screen "Proses" 800x480, template "Template_1"
   TextField "Text field_18" at 473,92 size 53x19; Text 'TT-0001'
   IOField "I/O field_11" at 473,110 size 55x20; FormatPattern 999; Unit  °C
      ProcessValue <- "TT-0001"
   TextField "Text field_19" at 548,92 size 53x19; Text 'TT-0002'
   IOField "I/O field_12" at 548,110 size 55x20; FormatPattern 999; Unit  °C
      ProcessValue <- "TT-0002"
   TextField "Text field_20" at 474,141 size 50x19; Text 'PT-0001'
   IOField "I/O field_13" at 474,159 size 52x20; FormatPattern 99; Unit  Bar
      ProcessValue <- "PT-0001"
   TextField "Text field_21" at 550,141 size 50x19; Text 'PT-0002'
   IOField "I/O field_14" at 550,159 size 52x20; FormatPattern 99; Unit  Bar
      ProcessValue <- "PT-0002"
   GraphicView "Graphic view_17" at 37,119 size 60x45; Picture "Graphic_29"
   Circle "Circle_3" at 95,98 size 16x16
      Appearance <- "PUMP_PUMP-1_Yedek1"
   TextField "Text field_67" at 24,118 size 16x22; Text 'R'
      Visibility <- "PUMP_PUMP-1_Local/Remote"
   TextField "Text field_68" at 26,119 size 14x22; Text 'L'
      Visibility <- "PUMP_PUMP-1_Local/Remote"
   TextField "Text field_10" at 28,97 size 49x20; Text 'PUMP-1'
   IOField "I/O field_15" at 71,167 size 45x20; FormatPattern 99; Unit  A
      ProcessValue <- "Pump-1_A"
   IOField "I/O field_6" at 24,167 size 45x20; FormatPattern 999; Unit  °C
      ProcessValue <- "Pump-1_Temp"
   GraphicView "Graphic view_1" at 145,119 size 60x45; Picture "Graphic_29"
   Circle "Circle_1" at 203,98 size 16x16
      Appearance <- "PUMP_PUMP-2_Yedek1"
   TextField "Text field_1" at 132,118 size 16x22; Text 'R'
      Visibility <- "PUMP_PUMP-2_Local/Remote"
   TextField "Text field_2" at 134,117 size 14x22; Text 'L'
      Visibility <- "PUMP_PUMP-2_Local/Remote"
   TextField "Text field_3" at 136,97 size 49x20; Text 'PUMP-2'
   IOField "I/O field_1" at 179,167 size 45x20; FormatPattern 99; Unit  A
      ProcessValue <- "Pump-2_A"
   IOField "I/O field_2" at 132,167 size 45x20; FormatPattern 999; Unit  °C
      ProcessValue <- "Pump-2_Temp"
   GraphicView "Graphic view_2" at 254,119 size 60x45; Picture "Graphic_29"
   Circle "Circle_2" at 312,98 size 16x16
      Appearance <- "PUMP_PUMP-3_Yedek1"
   TextField "Text field_4" at 241,118 size 16x22; Text 'R'
      Visibility <- "PUMP_PUMP-3_Local/Remote"
   TextField "Text field_5" at 243,117 size 14x22; Text 'L'
      Visibility <- "PUMP_PUMP-3_Local/Remote"
   TextField "Text field_6" at 245,97 size 49x20; Text 'PUMP-3'
   IOField "I/O field_3" at 288,167 size 45x20; FormatPattern 99; Unit  A
      ProcessValue <- "Pump-3_A"
   IOField "I/O field_4" at 241,167 size 45x20; FormatPattern 999; Unit  °C
      ProcessValue <- "Pump-3_Temp"
   GraphicView "Graphic view_3" at 360,119 size 60x45; Picture "Graphic_29"
   Circle "Circle_4" at 418,98 size 16x16
      Appearance <- "PUMP_PUMP-4_Yedek1"
   TextField "Text field_7" at 347,118 size 16x22; Text 'R'
      Visibility <- "PUMP_PUMP-4_Local/Remote"
   TextField "Text field_8" at 349,117 size 14x22; Text 'L'
      Visibility <- "PUMP_PUMP-4_Local/Remote"
   TextField "Text field_9" at 351,97 size 49x20; Text 'PUMP-4'
   IOField "I/O field_5" at 394,167 size 45x20; FormatPattern 99; Unit  A
      ProcessValue <- "Pump-4_A"
   IOField "I/O field_7" at 347,167 size 45x20; FormatPattern 999; Unit  °C
      ProcessValue <- "Pump-4_Temp"
   IOField "I/O field_22" at 40,269 size 51x20; FormatPattern 9999; Unit  %
      ProcessValue <- "CValve-1_Fbk"
   TextField "Text field_70" at 32,212 size 74x19; Text 'CONTROL V-1'
   GraphicView "Template_Graphic view_5" at 44,232 size 38x32; Picture "Graphic_74"
   IOField "I/O field_8" at 148,269 size 51x20; FormatPattern 9999; Unit  %
      ProcessValue <- "CValve-2_Fbk"
   GraphicView "Template_Graphic view_1" at 152,232 size 38x32; Picture "Graphic_74"
   TextField "Text field_12" at 140,212 size 74x19; Text 'CONTROL V-2'
   IOField "I/O field_9" at 257,269 size 51x20; FormatPattern 9999; Unit  %
      ProcessValue <- "CValve-3_Fbk"
   GraphicView "Template_Graphic view_2" at 261,232 size 38x32; Picture "Graphic_74"
   TextField "Text field_14" at 248,212 size 74x19; Text 'CONTROL V-3'
   IOField "I/O field_10" at 363,269 size 51x20; FormatPattern 9999; Unit  %
      ProcessValue <- "CValve-4_Fbk"
   GraphicView "Template_Graphic view_3" at 367,232 size 38x32; Picture "Graphic_74"
   TextField "Text field_16" at 354,212 size 74x19; Text 'CONTROL V-4'
   TextField "Text field_22" at 55,320 size 47x19; Text 'VALVE-1'
   Circle "Circle_23" at 37,322 size 16x16
      Appearance <- "VALVE-H_VALVE-1_ValveStatus"
   GraphicView "Graphic view_5" at 56,343 size 35x33; Picture "Graphic_102"
   TextField "Text field_23" at 160,320 size 47x19; Text 'VALVE-2'
   Circle "Circle_5" at 142,322 size 16x16
      Appearance <- "VALVE-H_VALVE-2_ValveStatus"
   GraphicView "Graphic view_4" at 161,343 size 35x33; Picture "Graphic_102"
   TextField "Text field_24" at 269,320 size 47x19; Text 'VALVE-3'
   Circle "Circle_6" at 251,322 size 16x16
      Appearance <- "VALVE-H_VALVE-3_ValveStatus"
   GraphicView "Graphic view_6" at 270,343 size 35x33; Picture "Graphic_102"
   TextField "Text field_25" at 375,320 size 47x19; Text 'VALVE-4'
   Circle "Circle_7" at 357,322 size 16x16
      Appearance <- "VALVE-H_VALVE-4_ValveStatus"
   GraphicView "Graphic view_7" at 376,343 size 35x33; Picture "Graphic_102"
   Button "Button_46" at 21,203 size 99x105; TextOff 'Text'
      on Press: InvertBit("HMI_Popup_POPUP{8}")
   Button "Button_1" at 127,203 size 99x105; TextOff 'Text'
      on Press: InvertBit("HMI_Popup_POPUP{9}")
   Button "Button_2" at 233,203 size 99x105; TextOff 'Text'
      on Press: InvertBit("HMI_Popup_POPUP{10}")
   Button "Button_3" at 339,210 size 99x98; TextOff 'Text'
      on Press: InvertBit("HMI_Popup_POPUP{11}")
   Button "Button_4" at 17,91 size 99x104; TextOff 'Text'
      on Press: InvertBit("HMI_Popup_POPUP{0}")
   Button "Button_5" at 126,92 size 99x103; TextOff 'Text'
      on Press: InvertBit("HMI_Popup_POPUP{1}")
   Button "Button_6" at 235,93 size 99x102; TextOff 'Text'
      on Press: InvertBit("HMI_Popup_POPUP{2}")
   Button "Button_7" at 344,86 size 99x108; TextOff 'Text'
      on Press: InvertBit("HMI_Popup_POPUP{3}")
   Button "Button_8" at 26,313 size 96x73; TextOff 'Text'
      on Press: InvertBit("HMI_Popup_POPUP{4}")
   Button "Button_9" at 129,313 size 95x72; TextOff 'Text'
      on Press: InvertBit("HMI_Popup_POPUP{5}")
   Button "Button_10" at 238,310 size 102x75; TextOff 'Text'
      on Press: InvertBit("HMI_Popup_POPUP{6}")
   Button "Button_11" at 348,314 size 95x72; TextOff 'Text'
      on Press: InvertBit("HMI_Popup_POPUP{7}")
   Group "Group" at 480,261 size 300x170
   Group "Group_1" at 480,261 size 300x170
   Group "Group_2" at 480,261 size 300x170
   Group "Group_3" at 480,261 size 300x170
   Group "Group_4" at 480,261 size 300x170
   Group "Group_5" at 480,261 size 300x170
   Group "Group_6" at 480,261 size 300x170
   Group "Group_7" at 480,261 size 300x170
   Group "Group_8" at 480,261 size 300x170
   Group "Group_9" at 480,261 size 300x170
   Group "Group_10" at 480,261 size 300x170
   Group "Group_11" at 480,261 size 300x170
   Rectangle "Rectangle_13" at 480,261 size 300x170
      Visibility <- "HMI_Popup_POPUP{4}"
   Button "Button_12" at 495,381 size 133x41; TextOn 'OPENED'; TextOff 'OPEN'
      on Release: ResetBit("VALVE-H_VALVE-1_ManuelOpen")
      on Press: SetBit("VALVE-H_VALVE-1_ManuelOpen")
      Visibility <- "HMI_Popup_POPUP{4}"
   Button "Button_13" at 633,381 size 133x41; TextOn 'CLOSED'; TextOff 'CLOSE'
      on Release: ResetBit("VALVE-H_VALVE-1_ManuelClose")
      on Press: SetBit("VALVE-H_VALVE-1_ManuelClose")
      Visibility <- "HMI_Popup_POPUP{4}"
   Switch "Switch_1" at 640,316 size 130x55; TextOn 'OTO'; CaptionText 'Switch'; TextOff 'MAN'
      Visibility <- "HMI_Popup_POPUP{4}"
   Button "Button_14" at 715,266 size 57x36; TextOff 'Text'; PictureOff "button"
      on Press: InvertBit("HMI_Popup_POPUP{4}")
      Visibility <- "HMI_Popup_POPUP{4}"
   TextField "Text field_11" at 490,271 size 134x33; Text 'VALVE-1'
      Visibility <- "HMI_Popup_POPUP{4}"
   Rectangle "Rectangle_14" at 575,336 size 20x18
      Visibility <- "HMI_Popup_POPUP{4}"
      Appearance <- "VALVE-H_VALVE-1_ValveStatus"
   TextField "Text field_13" at 502,336 size 45x17; Text 'OPENED'
      Visibility <- "HMI_Popup_POPUP{4}"
   Rectangle "Rectangle_15" at 480,261 size 300x170
      Visibility <- "HMI_Popup_POPUP{5}"
   Button "Button_15" at 495,381 size 133x41; TextOn 'OPENED'; TextOff 'OPEN'
      on Release: ResetBit("VALVE-H_VALVE-2_ManuelOpen")
      on Press: SetBit("VALVE-H_VALVE-2_ManuelOpen")
      Visibility <- "HMI_Popup_POPUP{5}"
   Button "Button_16" at 633,381 size 133x41; TextOn 'CLOSED'; TextOff 'CLOSE'
      on Release: ResetBit("VALVE-H_VALVE-2_ManuelClose")
      on Press: SetBit("VALVE-H_VALVE-2_ManuelClose")
      Visibility <- "HMI_Popup_POPUP{5}"
   Switch "Switch_2" at 640,316 size 130x55; TextOn 'OTO'; CaptionText 'Switch'; TextOff 'MAN'
      Visibility <- "HMI_Popup_POPUP{5}"
   Button "Button_17" at 715,266 size 57x36; TextOff 'Text'; PictureOff "button"
      on Press: InvertBit("HMI_Popup_POPUP{5}")
      Visibility <- "HMI_Popup_POPUP{5}"
   TextField "Text field_15" at 490,271 size 134x33; Text 'VALVE-2'
      Visibility <- "HMI_Popup_POPUP{5}"
   Rectangle "Rectangle_16" at 575,336 size 20x18
      Visibility <- "HMI_Popup_POPUP{5}"
      Appearance <- "VALVE-H_VALVE-2_ValveStatus"
   TextField "Text field_17" at 502,336 size 45x17; Text 'OPENED'
      Visibility <- "HMI_Popup_POPUP{5}"
   Rectangle "Rectangle_17" at 480,261 size 300x170
      Visibility <- "HMI_Popup_POPUP{7}"
   Button "Button_18" at 495,381 size 133x41; TextOn 'OPENED'; TextOff 'OPEN'
      on Release: ResetBit("VALVE-H_VALVE-4_ManuelOpen")
      on Press: SetBit("VALVE-H_VALVE-4_ManuelOpen")
      Visibility <- "HMI_Popup_POPUP{7}"
   Button "Button_19" at 633,381 size 133x41; TextOn 'CLOSED'; TextOff 'CLOSE'
      on Release: ResetBit("VALVE-H_VALVE-4_ManuelClose")
      on Press: SetBit("VALVE-H_VALVE-4_ManuelClose")
      Visibility <- "HMI_Popup_POPUP{7}"
   Switch "Switch_4" at 640,316 size 130x55; TextOn 'OTO'; CaptionText 'Switch'; TextOff 'MAN'
      Visibility <- "HMI_Popup_POPUP{7}"
   Button "Button_20" at 715,266 size 57x36; TextOff 'Text'; PictureOff "button"
      on Press: InvertBit("HMI_Popup_POPUP{7}")
      Visibility <- "HMI_Popup_POPUP{7}"
   TextField "Text field_26" at 490,271 size 134x33; Text 'VALVE-4'
      Visibility <- "HMI_Popup_POPUP{7}"
   Rectangle "Rectangle_18" at 575,336 size 20x18
      Visibility <- "HMI_Popup_POPUP{7}"
      Appearance <- "VALVE-H_VALVE-4_ValveStatus"
   TextField "Text field_27" at 502,336 size 45x17; Text 'OPENED'
      Visibility <- "HMI_Popup_POPUP{7}"
   Rectangle "Rectangle_19" at 480,261 size 300x170
      Visibility <- "HMI_Popup_POPUP{6}"
   Button "Button_21" at 495,381 size 133x41; TextOn 'OPENED'; TextOff 'OPEN'
      on Release: ResetBit("VALVE-H_VALVE-3_ManuelOpen")
      on Press: SetBit("VALVE-H_VALVE-3_ManuelOpen")
      Visibility <- "HMI_Popup_POPUP{6}"
   Button "Button_22" at 633,381 size 133x41; TextOn 'CLOSED'; TextOff 'CLOSE'
      on Release: ResetBit("VALVE-H_VALVE-3_ManuelClose")
      on Press: SetBit("VALVE-H_VALVE-3_ManuelClose")
      Visibility <- "HMI_Popup_POPUP{6}"
   Switch "Switch_3" at 640,316 size 130x55; TextOn 'OTO'; CaptionText 'Switch'; TextOff 'MAN'
      Visibility <- "HMI_Popup_POPUP{6}"
   Button "Button_23" at 715,266 size 57x36; TextOff 'Text'; PictureOff "button"
      on Press: InvertBit("HMI_Popup_POPUP{6}")
      Visibility <- "HMI_Popup_POPUP{6}"
   TextField "Text field_28" at 490,271 size 134x33; Text 'VALVE-3'
      Visibility <- "HMI_Popup_POPUP{6}"
   Rectangle "Rectangle_20" at 575,336 size 20x18
      Visibility <- "HMI_Popup_POPUP{6}"
      Appearance <- "VALVE-H_VALVE-3_ValveStatus"
   TextField "Text field_29" at 502,336 size 45x17; Text 'OPENED'
      Visibility <- "HMI_Popup_POPUP{6}"
   Rectangle "Rectangle_21" at 480,261 size 300x170
      Visibility <- "HMI_Popup_POPUP{0}"
   Button "Button_47" at 637,368 size 130x40; TextOn 'STOPPED'; TextOff 'STOP'
      on Release: ResetBit("PUMP_PUMP-1_ManuelStop")
      on Press: SetBit("PUMP_PUMP-1_ManuelStop")
      Visibility <- "HMI_Popup_POPUP{0}"
   Button "Button_48" at 636,317 size 130x40; TextOn 'STARTED'; TextOff 'START'
      on Release: ResetBit("PUMP_PUMP-1_ManuelStart")
      on Press: SetBit("PUMP_PUMP-1_ManuelStart")
      Visibility <- "HMI_Popup_POPUP{0}"
   IOField "I/O field_16" at 509,391 size 106x35; FormatPattern 9999; Unit    Rpm
      ProcessValue <- "HMI_Pump-1"
      Visibility <- "HMI_Popup_POPUP{0}"
   Button "Button_49" at 715,268 size 57x36; TextOff 'Text'; PictureOff "button"
      on Press: InvertBit("HMI_Popup_POPUP{0}")
      Visibility <- "HMI_Popup_POPUP{0}"
   TextField "Text field_64" at 503,270 size 86x33; Text 'PUMP-1'
      Visibility <- "HMI_Popup_POPUP{0}"
   Rectangle "Rectangle_22" at 572,334 size 20x18
      Visibility <- "HMI_Popup_POPUP{0}"
      Appearance <- "PUMP_PUMP-1_MotorStatus"
   Rectangle "Rectangle_23" at 572,312 size 20x18
      Visibility <- "HMI_Popup_POPUP{0}"
      Appearance <- "PUMP_PUMP-1_MotorStatus"
   Rectangle "Rectangle_24" at 572,356 size 20x18
      Visibility <- "HMI_Popup_POPUP{0}"
      Appearance <- "PUMP_PUMP-1_MotorStatus"
   TextField "Text field_30" at 498,314 size 51x17; Text 'RUNNING'
      Visibility <- "HMI_Popup_POPUP{0}"
   TextField "Text field_33" at 499,333 size 61x17; Text 'INTERLOCK'
      Visibility <- "HMI_Popup_POPUP{0}"
   TextField "Text field_34" at 499,353 size 36x17; Text 'FAULT'
      Visibility <- "HMI_Popup_POPUP{0}"
   Rectangle "Rectangle_25" at 480,261 size 300x170
      Visibility <- "HMI_Popup_POPUP{1}"
   Button "Button_24" at 637,368 size 130x40; TextOn 'STOPPED'; TextOff 'STOP'
      on Release: ResetBit("PUMP_PUMP-2_ManuelStop")
      on Press: SetBit("PUMP_PUMP-2_ManuelStop")
      Visibility <- "HMI_Popup_POPUP{1}"
   Button "Button_25" at 636,317 size 130x40; TextOn 'STARTED'; TextOff 'START'
      on Release: ResetBit("PUMP_PUMP-2_ManuelStart")
      on Press: SetBit("PUMP_PUMP-2_ManuelStart")
      Visibility <- "HMI_Popup_POPUP{1}"
   IOField "I/O field_17" at 509,391 size 106x35; FormatPattern 9999; Unit    Rpm
      ProcessValue <- "HMI_Pump-2"
      Visibility <- "HMI_Popup_POPUP{1}"
   Button "Button_26" at 715,268 size 57x36; TextOff 'Text'; PictureOff "button"
      on Press: InvertBit("HMI_Popup_POPUP{1}")
      Visibility <- "HMI_Popup_POPUP{1}"
   TextField "Text field_31" at 503,270 size 86x33; Text 'PUMP-2'
      Visibility <- "HMI_Popup_POPUP{1}"
   Rectangle "Rectangle_26" at 572,334 size 20x18
      Visibility <- "HMI_Popup_POPUP{1}"
      Appearance <- "PUMP_PUMP-2_MotorStatus"
   Rectangle "Rectangle_27" at 572,312 size 20x18
      Visibility <- "HMI_Popup_POPUP{1}"
      Appearance <- "PUMP_PUMP-2_MotorStatus"
   Rectangle "Rectangle_28" at 572,356 size 20x18
      Visibility <- "HMI_Popup_POPUP{1}"
      Appearance <- "PUMP_PUMP-2_MotorStatus"
   TextField "Text field_32" at 498,314 size 51x17; Text 'RUNNING'
      Visibility <- "HMI_Popup_POPUP{1}"
   TextField "Text field_35" at 499,333 size 61x17; Text 'INTERLOCK'
      Visibility <- "HMI_Popup_POPUP{1}"
   TextField "Text field_36" at 499,353 size 36x17; Text 'FAULT'
      Visibility <- "HMI_Popup_POPUP{1}"
   Rectangle "Rectangle_29" at 480,261 size 300x170
      Visibility <- "HMI_Popup_POPUP{3}"
   Button "Button_27" at 637,368 size 130x40; TextOn 'STOPPED'; TextOff 'STOP'
      on Release: ResetBit("PUMP_PUMP-4_ManuelStop")
      on Press: SetBit("PUMP_PUMP-4_ManuelStop")
      Visibility <- "HMI_Popup_POPUP{3}"
   Button "Button_28" at 636,317 size 130x40; TextOn 'STARTED'; TextOff 'START'
      on Release: ResetBit("PUMP_PUMP-4_ManuelStart")
      on Press: SetBit("PUMP_PUMP-4_ManuelStart")
      Visibility <- "HMI_Popup_POPUP{3}"
   IOField "I/O field_18" at 509,391 size 106x35; FormatPattern 9999; Unit    Rpm
      ProcessValue <- "HMI_Pump-4"
      Visibility <- "HMI_Popup_POPUP{3}"
   Button "Button_29" at 715,268 size 57x36; TextOff 'Text'; PictureOff "button"
      on Press: InvertBit("HMI_Popup_POPUP{3}")
      Visibility <- "HMI_Popup_POPUP{3}"
   TextField "Text field_37" at 503,270 size 86x33; Text 'PUMP-4'
      Visibility <- "HMI_Popup_POPUP{3}"
   Rectangle "Rectangle_30" at 572,334 size 20x18
      Visibility <- "HMI_Popup_POPUP{3}"
      Appearance <- "PUMP_PUMP-4_MotorStatus"
   Rectangle "Rectangle_31" at 572,312 size 20x18
      Visibility <- "HMI_Popup_POPUP{3}"
      Appearance <- "PUMP_PUMP-4_MotorStatus"
   Rectangle "Rectangle_32" at 572,356 size 20x18
      Visibility <- "HMI_Popup_POPUP{3}"
      Appearance <- "PUMP_PUMP-4_MotorStatus"
   TextField "Text field_38" at 498,314 size 51x17; Text 'RUNNING'
      Visibility <- "HMI_Popup_POPUP{3}"
   TextField "Text field_39" at 499,333 size 61x17; Text 'INTERLOCK'
      Visibility <- "HMI_Popup_POPUP{3}"
   TextField "Text field_40" at 499,353 size 36x17; Text 'FAULT'
      Visibility <- "HMI_Popup_POPUP{3}"
   Rectangle "Rectangle_33" at 480,261 size 300x170
      Visibility <- "HMI_Popup_POPUP{2}"
   Button "Button_30" at 637,368 size 130x40; TextOn 'STOPPED'; TextOff 'STOP'
      on Release: ResetBit("PUMP_PUMP-3_ManuelStop")
      on Press: SetBit("PUMP_PUMP-3_ManuelStop")
      Visibility <- "HMI_Popup_POPUP{2}"
   Button "Button_31" at 636,317 size 130x40; TextOn 'STARTED'; TextOff 'START'
      on Release: ResetBit("PUMP_PUMP-3_ManuelStart")
      on Press: SetBit("PUMP_PUMP-3_ManuelStart")
      Visibility <- "HMI_Popup_POPUP{2}"
   IOField "I/O field_19" at 509,391 size 106x35; FormatPattern 9999; Unit    Rpm
      ProcessValue <- "HMI_Pump-3"
      Visibility <- "HMI_Popup_POPUP{2}"
   Button "Button_32" at 715,268 size 57x36; TextOff 'Text'; PictureOff "button"
      on Press: InvertBit("HMI_Popup_POPUP{2}")
      Visibility <- "HMI_Popup_POPUP{2}"
   TextField "Text field_41" at 503,270 size 86x33; Text 'PUMP-3'
      Visibility <- "HMI_Popup_POPUP{2}"
   Rectangle "Rectangle_34" at 572,334 size 20x18
      Visibility <- "HMI_Popup_POPUP{2}"
      Appearance <- "PUMP_PUMP-3_MotorStatus"
   Rectangle "Rectangle_35" at 572,312 size 20x18
      Visibility <- "HMI_Popup_POPUP{2}"
      Appearance <- "PUMP_PUMP-3_MotorStatus"
   Rectangle "Rectangle_36" at 572,356 size 20x18
      Visibility <- "HMI_Popup_POPUP{2}"
      Appearance <- "PUMP_PUMP-3_MotorStatus"
   TextField "Text field_42" at 498,314 size 51x17; Text 'RUNNING'
      Visibility <- "HMI_Popup_POPUP{2}"
   TextField "Text field_43" at 499,333 size 61x17; Text 'INTERLOCK'
      Visibility <- "HMI_Popup_POPUP{2}"
   TextField "Text field_44" at 499,353 size 36x17; Text 'FAULT'
      Visibility <- "HMI_Popup_POPUP{2}"
   Rectangle "Rectangle_37" at 480,261 size 300x170
      Visibility <- "HMI_Popup_POPUP{8}"
   IOField "I/O field_20" at 503,355 size 101x35; FormatPattern 999; Unit  %
      ProcessValue <- "HMI_CValve-1_Set"
      Visibility <- "HMI_Popup_POPUP{8}"
   TextField "Text field_45" at 487,271 size 175x32; Text 'CONTROL VALVE-1'
      Visibility <- "HMI_Popup_POPUP{8}"
   Switch "Switch_5" at 631,343 size 130x55; TextOn 'OTO'; CaptionText 'Switch'; TextOff 'MAN'
      Visibility <- "HMI_Popup_POPUP{8}"
   Button "Button_33" at 716,268 size 57x36; TextOff 'Text'; PictureOff "button"
      on Press: InvertBit("HMI_Popup_POPUP{8}")
      Visibility <- "HMI_Popup_POPUP{8}"
   Rectangle "Rectangle_38" at 480,261 size 300x170
      Visibility <- "HMI_Popup_POPUP{9}"
   IOField "I/O field_21" at 503,355 size 101x35; FormatPattern 999; Unit  %
      ProcessValue <- "HMI_CValve-2_Set"
      Visibility <- "HMI_Popup_POPUP{9}"
   TextField "Text field_46" at 487,271 size 175x32; Text 'CONTROL VALVE-2'
      Visibility <- "HMI_Popup_POPUP{9}"
   Switch "Switch_6" at 631,343 size 130x55; TextOn 'OTO'; CaptionText 'Switch'; TextOff 'MAN'
      Visibility <- "HMI_Popup_POPUP{9}"
   Button "Button_34" at 716,268 size 57x36; TextOff 'Text'; PictureOff "button"
      on Press: InvertBit("HMI_Popup_POPUP{9}")
      Visibility <- "HMI_Popup_POPUP{9}"
   Rectangle "Rectangle_39" at 480,261 size 300x170
      Visibility <- "HMI_Popup_POPUP{11}"
   IOField "I/O field_23" at 503,355 size 101x35; FormatPattern 999; Unit  %
      Visibility <- "HMI_Popup_POPUP{11}"
      ProcessValue <- "HMI_CValve-4_Set"
   TextField "Text field_47" at 487,271 size 175x32; Text 'CONTROL VALVE-4'
      Visibility <- "HMI_Popup_POPUP{11}"
   Switch "Switch_7" at 631,343 size 130x55; TextOn 'OTO'; CaptionText 'Switch'; TextOff 'MAN'
      Visibility <- "HMI_Popup_POPUP{11}"
   Button "Button_35" at 716,268 size 57x36; TextOff 'Text'; PictureOff "button"
      on Press: InvertBit("HMI_Popup_POPUP{11}")
      Visibility <- "HMI_Popup_POPUP{11}"
   Rectangle "Rectangle_40" at 480,261 size 300x170
      Visibility <- "HMI_Popup_POPUP{10}"
   IOField "I/O field_24" at 503,355 size 101x35; FormatPattern 999; Unit  %
      ProcessValue <- "HMI_CValve-3_Set"
      Visibility <- "HMI_Popup_POPUP{10}"
   TextField "Text field_48" at 487,271 size 175x32; Text 'CONTROL VALVE-3'
      Visibility <- "HMI_Popup_POPUP{10}"
   Switch "Switch_8" at 631,343 size 130x55; TextOn 'OTO'; CaptionText 'Switch'; TextOff 'MAN'
      Visibility <- "HMI_Popup_POPUP{10}"
   Button "Button_36" at 716,268 size 57x36; TextOff 'Text'; PictureOff "button"
      on Press: InvertBit("HMI_Popup_POPUP{10}")
      Visibility <- "HMI_Popup_POPUP{10}"

screen "Con" 800x480, template "Template_1"
   TextField "Text field_8" at 56,79 size 84x20; Text 'Work Order-1'
   TextField "Text field_13" at 352,163 size 124x20; Text 'Work Order Select'
   TextField "Text field_14" at 593,165 size 118x20; Text 'Work Order Start'
   TextField "Text field_1" at 56,102 size 84x20; Text 'Work Order-2'
   TextField "Text field_2" at 56,125 size 84x20; Text 'Work Order-3'
   TextField "Text field_3" at 56,148 size 84x20; Text 'Work Order-4'
   TextField "Text field_4" at 56,171 size 84x20; Text 'Work Order-5'
   TextField "Text field_5" at 56,195 size 84x20; Text 'Work Order-6'
   TextField "Text field_6" at 56,218 size 84x20; Text 'Work Order-7'
   TextField "Text field_7" at 56,241 size 84x20; Text 'Work Order-8'
   TextField "Text field_9" at 56,264 size 84x20; Text 'Work Order-9'
   TextField "Text field_10" at 56,288 size 91x20; Text 'Work Order-10'
   TextField "Text field_16" at 56,312 size 91x20; Text 'Work Order-11'
   TextField "Text field_17" at 56,335 size 91x20; Text 'Work Order-12'
   TextField "Text field_18" at 56,359 size 91x20; Text 'Work Order-13'
   TextField "Text field_19" at 56,383 size 91x20; Text 'Work Order-14'
   TextField "Text field_11" at 222,77 size 51x20; Text 'ACTIVE'
      Visibility <- "workorder_Work_Order-1_Active"
   TextField "Text field_20" at 213,77 size 60x20; Text 'PASSIVE'
      Visibility <- "workorder_Work_Order-1_Active"
   TextField "Text field_21" at 222,100 size 51x20; Text 'ACTIVE'
      Visibility <- "workorder_Work_Order-2_Active"
   TextField "Text field_22" at 222,123 size 51x20; Text 'ACTIVE'
      Visibility <- "workorder_Work_Order-3_Active"
   TextField "Text field_23" at 222,147 size 51x20; Text 'ACTIVE'
      Visibility <- "workorder_Work_Order-4_Active"
   TextField "Text field_24" at 222,170 size 51x21; Text 'ACTIVE'
      Visibility <- "workorder_Work_Order-5_Active"
   TextField "Text field_25" at 222,195 size 51x20; Text 'ACTIVE'
      Visibility <- "workorder_Work_Order-6_Active"
   TextField "Text field_26" at 222,218 size 51x21; Text 'ACTIVE'
      Visibility <- "workorder_Work_Order-7_Active"
   TextField "Text field_27" at 222,243 size 51x20; Text 'ACTIVE'
      Visibility <- "workorder_Work_Order-8_Active"
   TextField "Text field_28" at 222,266 size 51x20; Text 'ACTIVE'
      Visibility <- "workorder_Work_Order-9_Active"
   TextField "Text field_29" at 222,290 size 51x20; Text 'ACTIVE'
      Visibility <- "workorder_Work_Order-10_Active"
   TextField "Text field_30" at 222,313 size 51x20; Text 'ACTIVE'
      Visibility <- "workorder_Work_Order-11_Active"
   TextField "Text field_31" at 222,337 size 51x20; Text 'ACTIVE'
      Visibility <- "workorder_Work_Order-12_Active"
   TextField "Text field_32" at 222,360 size 51x20; Text 'ACTIVE'
      Visibility <- "workorder_Work_Order-13_Active"
   TextField "Text field_33" at 222,384 size 51x21; Text 'ACTIVE'
      Visibility <- "workorder_Work_Order-14_Active"
   TextField "Text field_34" at 213,100 size 60x20; Text 'PASSIVE'
      Visibility <- "workorder_Work_Order-2_Active"
   TextField "Text field_35" at 213,124 size 60x20; Text 'PASSIVE'
      Visibility <- "workorder_Work_Order-3_Active"
   TextField "Text field_36" at 213,147 size 60x20; Text 'PASSIVE'
      Visibility <- "workorder_Work_Order-4_Active"
   TextField "Text field_37" at 213,171 size 60x20; Text 'PASSIVE'
      Visibility <- "workorder_Work_Order-5_Active"
   TextField "Text field_38" at 213,194 size 60x21; Text 'PASSIVE'
      Visibility <- "workorder_Work_Order-6_Active"
   TextField "Text field_39" at 213,219 size 60x20; Text 'PASSIVE'
      Visibility <- "workorder_Work_Order-7_Active"
   TextField "Text field_40" at 213,242 size 60x20; Text 'PASSIVE'
      Visibility <- "workorder_Work_Order-8_Active"
   TextField "Text field_41" at 213,266 size 60x20; Text 'PASSIVE'
      Visibility <- "workorder_Work_Order-9_Active"
   TextField "Text field_42" at 213,289 size 60x20; Text 'PASSIVE'
      Visibility <- "workorder_Work_Order-10_Active"
   TextField "Text field_43" at 213,313 size 60x20; Text 'PASSIVE'
      Visibility <- "workorder_Work_Order-11_Active"
   TextField "Text field_44" at 213,336 size 60x20; Text 'PASSIVE'
      Visibility <- "workorder_Work_Order-12_Active"
   TextField "Text field_45" at 213,360 size 60x20; Text 'PASSIVE'
      Visibility <- "workorder_Work_Order-13_Active"
   TextField "Text field_46" at 213,384 size 60x21; Text 'PASSIVE'
      Visibility <- "workorder_Work_Order-14_Active"
   SymbolicIOField "Symbolic I/O field_1" at 344,216 size 156x32; TextOff '0'; TextOn '1'; TextList "WorkOrder"
   Button "Button_1" at 577,218 size 140x32; TextOff 'START'

screen "popup_motor" 800x480
   Rectangle "Rectangle_21" at 30,21 size 300x170
      Visibility <- "HMI_Popup_POPUP{0}"
   Button "Button_47" at 187,128 size 130x40; TextOn 'DURDU'; TextOff 'STOP'
      on Release: ResetBit("PUMP_PUMP-1_ManuelStop")
      on Press: SetBit("PUMP_PUMP-1_ManuelStop")
      Visibility <- "HMI_Popup_POPUP{0}"
   Button "Button_48" at 186,77 size 130x40; TextOn 'ÇALIŞTI'; TextOff 'START'
      on Release: ResetBit("PUMP_PUMP-1_ManuelStart")
      on Press: SetBit("PUMP_PUMP-1_ManuelStart")
      Visibility <- "HMI_Popup_POPUP{0}"
   IOField "I/O field_14" at 59,151 size 106x35; FormatPattern 9999; Unit    Rpm
      Visibility <- "HMI_Popup_POPUP{0}"
      ProcessValue <- "HMI_Pump-1"
   Button "Button_49" at 265,28 size 57x36; TextOff 'Text'; PictureOff "button"
      on Press: InvertBit("HMI_Popup_POPUP{0}")
      Visibility <- "HMI_Popup_POPUP{0}"
   TextField "Text field_64" at 53,30 size 86x33; Text 'PUMP-1'
      Visibility <- "HMI_Popup_POPUP{0}"
   Rectangle "Rectangle_14" at 122,94 size 20x18
      Visibility <- "HMI_Popup_POPUP{0}"
      Appearance <- "PUMP_PUMP-1_MotorStatus"
   Rectangle "Rectangle_16" at 122,72 size 20x18
      Visibility <- "HMI_Popup_POPUP{0}"
      Appearance <- "PUMP_PUMP-1_MotorStatus"
   Rectangle "Rectangle_22" at 122,116 size 20x18
      Visibility <- "HMI_Popup_POPUP{0}"
      Appearance <- "PUMP_PUMP-1_MotorStatus"
   TextField "Text field_30" at 48,74 size 51x17; Text 'RUNNING'
      Visibility <- "HMI_Popup_POPUP{0}"
   TextField "Text field_33" at 49,93 size 61x17; Text 'INTERLOCK'
      Visibility <- "HMI_Popup_POPUP{0}"
   TextField "Text field_34" at 49,113 size 36x17; Text 'FAULT'
      Visibility <- "HMI_Popup_POPUP{0}"
   Rectangle "Rectangle_5" at 37,222 size 300x170
      Visibility <- "HMI_Popup_POPUP{2}"
   Button "Button_4" at 194,329 size 130x40; TextOn 'DURDU'; TextOff 'STOP'
      on Release: ResetBit("PUMP_PUMP-3_ManuelStop")
      on Press: SetBit("PUMP_PUMP-3_ManuelStop")
      Visibility <- "HMI_Popup_POPUP{2}"
   Button "Button_5" at 193,278 size 130x40; TextOn 'ÇALIŞTI'; TextOff 'START'
      on Release: ResetBit("PUMP_PUMP-3_ManuelStart")
      on Press: SetBit("PUMP_PUMP-3_ManuelStart")
      Visibility <- "HMI_Popup_POPUP{2}"
   IOField "I/O field_2" at 66,352 size 106x35; FormatPattern 9999; Unit    Rpm
      Visibility <- "HMI_Popup_POPUP{2}"
      ProcessValue <- "HMI_Pump-3"
   Button "Button_6" at 272,229 size 57x36; TextOff 'Text'; PictureOff "button"
      on Press: InvertBit("HMI_Popup_POPUP{2}")
      Visibility <- "HMI_Popup_POPUP{2}"
   TextField "Text field_5" at 60,231 size 86x33; Text 'PUMP-3'
      Visibility <- "HMI_Popup_POPUP{2}"
   Rectangle "Rectangle_6" at 129,295 size 20x18
      Visibility <- "HMI_Popup_POPUP{2}"
      Appearance <- "PUMP_PUMP-3_MotorStatus"
   Rectangle "Rectangle_7" at 129,273 size 20x18
      Visibility <- "HMI_Popup_POPUP{2}"
      Appearance <- "PUMP_PUMP-3_MotorStatus"
   Rectangle "Rectangle_8" at 129,317 size 20x18
      Visibility <- "HMI_Popup_POPUP{2}"
      Appearance <- "PUMP_PUMP-3_MotorStatus"
   TextField "Text field_6" at 55,275 size 51x17; Text 'RUNNING'
      Visibility <- "HMI_Popup_POPUP{2}"
   TextField "Text field_7" at 56,294 size 61x17; Text 'INTERLOCK'
      Visibility <- "HMI_Popup_POPUP{2}"
   TextField "Text field_8" at 56,314 size 36x17; Text 'FAULT'
      Visibility <- "HMI_Popup_POPUP{2}"
   Rectangle "Rectangle_9" at 384,217 size 300x170
      Visibility <- "HMI_Popup_POPUP{3}"
   Button "Button_7" at 541,324 size 130x40; TextOn 'DURDU'; TextOff 'STOP'
      on Release: ResetBit("PUMP_PUMP-4_ManuelStop")
      on Press: SetBit("PUMP_PUMP-4_ManuelStop")
      Visibility <- "HMI_Popup_POPUP{3}"
   Button "Button_8" at 540,273 size 130x40; TextOn 'ÇALIŞTI'; TextOff 'START'
      on Release: ResetBit("PUMP_PUMP-4_ManuelStart")
      on Press: SetBit("PUMP_PUMP-4_ManuelStart")
      Visibility <- "HMI_Popup_POPUP{3}"
   IOField "I/O field_3" at 413,347 size 106x35; FormatPattern 9999; Unit    Rpm
      Visibility <- "HMI_Popup_POPUP{3}"
      ProcessValue <- "HMI_Pump-4"
   Button "Button_9" at 619,224 size 57x36; TextOff 'Text'; PictureOff "button"
      on Press: InvertBit("HMI_Popup_POPUP{3}")
      Visibility <- "HMI_Popup_POPUP{3}"
   TextField "Text field_9" at 407,226 size 86x33; Text 'PUMP-4'
      Visibility <- "HMI_Popup_POPUP{3}"
   Rectangle "Rectangle_10" at 476,290 size 20x18
      Visibility <- "HMI_Popup_POPUP{3}"
      Appearance <- "PUMP_PUMP-4_MotorStatus"
   Rectangle "Rectangle_11" at 476,268 size 20x18
      Visibility <- "HMI_Popup_POPUP{3}"
      Appearance <- "PUMP_PUMP-4_MotorStatus"
   Rectangle "Rectangle_12" at 476,312 size 20x18
      Visibility <- "HMI_Popup_POPUP{3}"
      Appearance <- "PUMP_PUMP-4_MotorStatus"
   TextField "Text field_10" at 402,270 size 51x17; Text 'RUNNING'
      Visibility <- "HMI_Popup_POPUP{3}"
   TextField "Text field_11" at 403,289 size 61x17; Text 'INTERLOCK'
      Visibility <- "HMI_Popup_POPUP{3}"
   TextField "Text field_12" at 403,309 size 36x17; Text 'FAULT'
      Visibility <- "HMI_Popup_POPUP{3}"
   Group "Group" at 30,21 size 300x170
   Group "Group_2" at 384,217 size 300x170
   Group "Group_3" at 37,222 size 300x170
   Rectangle "Rectangle_1" at 383,21 size 300x170
      Visibility <- "HMI_Popup_POPUP{1}"
   Button "Button_1" at 540,128 size 130x40; TextOn 'DURDU'; TextOff 'STOP'
      on Release: ResetBit("PUMP_PUMP-2_ManuelStop")
      on Press: SetBit("PUMP_PUMP-2_ManuelStop")
      Visibility <- "HMI_Popup_POPUP{1}"
   Button "Button_2" at 539,77 size 130x40; TextOn 'ÇALIŞTI'; TextOff 'START'
      on Release: ResetBit("PUMP_PUMP-2_ManuelStart")
      on Press: SetBit("PUMP_PUMP-2_ManuelStart")
      Visibility <- "HMI_Popup_POPUP{1}"
   IOField "I/O field_1" at 412,151 size 106x35; FormatPattern 9999; Unit    Rpm
      Visibility <- "HMI_Popup_POPUP{1}"
      ProcessValue <- "HMI_Pump-2"
   Button "Button_3" at 618,28 size 57x36; TextOff 'Text'; PictureOff "button"
      on Press: InvertBit("HMI_Popup_POPUP{1}")
      Visibility <- "HMI_Popup_POPUP{1}"
   TextField "Text field_1" at 406,30 size 86x33; Text 'PUMP-2'
      Visibility <- "HMI_Popup_POPUP{1}"
   Rectangle "Rectangle_2" at 475,94 size 20x18
      Visibility <- "HMI_Popup_POPUP{1}"
      Appearance <- "PUMP_PUMP-2_MotorStatus"
   Rectangle "Rectangle_3" at 475,72 size 20x18
      Visibility <- "HMI_Popup_POPUP{1}"
      Appearance <- "PUMP_PUMP-2_MotorStatus"
   Rectangle "Rectangle_4" at 475,116 size 20x18
      Visibility <- "HMI_Popup_POPUP{1}"
      Appearance <- "PUMP_PUMP-2_MotorStatus"
   TextField "Text field_2" at 401,74 size 51x17; Text 'RUNNING'
      Visibility <- "HMI_Popup_POPUP{1}"
   TextField "Text field_3" at 402,93 size 61x17; Text 'INTERLOCK'
      Visibility <- "HMI_Popup_POPUP{1}"
   TextField "Text field_4" at 402,113 size 36x17; Text 'FAULT'
      Visibility <- "HMI_Popup_POPUP{1}"

screen "popup_vana" 800x480
   Rectangle "Rectangle_1" at 20,20 size 300x170
      Visibility <- "HMI_Popup_POPUP{4}"
   Button "Button_1" at 35,140 size 133x41; TextOn 'AÇILDI'; TextOff 'OPEN'
      on Press: SetBit("VALVE-H_VALVE-1_ManuelOpen")
      Visibility <- "HMI_Popup_POPUP{4}"
      on Release: ResetBit("VALVE-H_VALVE-1_ManuelOpen")
   Button "Button_2" at 173,140 size 133x41; TextOn 'KAPANDI'; TextOff 'CLOSE'
      on Press: SetBit("VALVE-H_VALVE-1_ManuelClose")
      Visibility <- "HMI_Popup_POPUP{4}"
      on Release: ResetBit("VALVE-H_VALVE-1_ManuelClose")
   Switch "Switch_1" at 180,75 size 130x55; TextOn 'OTO'; CaptionText 'Switch'; TextOff 'MAN'
      Visibility <- "HMI_Popup_POPUP{4}"
   Button "Button_3" at 255,25 size 57x36; TextOff 'Text'; PictureOff "button"
      on Press: InvertBit("HMI_Popup_POPUP{4}")
      Visibility <- "HMI_Popup_POPUP{4}"
   TextField "Text field_1" at 30,30 size 134x33; Text 'VALVE-1'
      Visibility <- "HMI_Popup_POPUP{4}"
   Rectangle "Rectangle_2" at 115,95 size 20x18
      Visibility <- "HMI_Popup_POPUP{4}"
      Appearance <- "VALVE-H_VALVE-1_ValveStatus"
   TextField "Text field_2" at 42,95 size 45x17; Text 'OPENED'
      Visibility <- "HMI_Popup_POPUP{4}"
   Rectangle "Rectangle_3" at 376,20 size 300x170
      Visibility <- "HMI_Popup_POPUP{5}"
   Button "Button_4" at 391,140 size 133x41; TextOn 'AÇILDI'; TextOff 'OPEN'
      on Press: SetBit("VALVE-H_VALVE-2_ManuelOpen")
      Visibility <- "HMI_Popup_POPUP{5}"
      on Release: ResetBit("VALVE-H_VALVE-2_ManuelOpen")
   Button "Button_5" at 529,140 size 133x41; TextOn 'KAPANDI'; TextOff 'CLOSE'
      on Press: SetBit("VALVE-H_VALVE-2_ManuelClose")
      Visibility <- "HMI_Popup_POPUP{5}"
      on Release: ResetBit("VALVE-H_VALVE-2_ManuelClose")
   Switch "Switch_2" at 536,75 size 130x55; TextOn 'OTO'; CaptionText 'Switch'; TextOff 'MAN'
      Visibility <- "HMI_Popup_POPUP{5}"
   Button "Button_6" at 611,25 size 57x36; TextOff 'Text'; PictureOff "button"
      on Press: InvertBit("HMI_Popup_POPUP{5}")
      Visibility <- "HMI_Popup_POPUP{5}"
   TextField "Text field_3" at 386,30 size 134x33; Text 'VALVE-2'
      Visibility <- "HMI_Popup_POPUP{5}"
   Rectangle "Rectangle_4" at 471,95 size 20x18
      Visibility <- "HMI_Popup_POPUP{5}"
      Appearance <- "VALVE-H_VALVE-2_ValveStatus"
   TextField "Text field_4" at 398,95 size 45x17; Text 'OPENED'
      Visibility <- "HMI_Popup_POPUP{5}"
   Rectangle "Rectangle_5" at 29,232 size 300x170
      Visibility <- "HMI_Popup_POPUP{6}"
   Button "Button_7" at 44,352 size 133x41; TextOn 'AÇILDI'; TextOff 'OPEN'
      on Press: SetBit("VALVE-H_VALVE-3_ManuelOpen")
      Visibility <- "HMI_Popup_POPUP{6}"
      on Release: ResetBit("VALVE-H_VALVE-3_ManuelOpen")
   Button "Button_8" at 182,352 size 133x41; TextOn 'KAPANDI'; TextOff 'CLOSE'
      on Press: SetBit("VALVE-H_VALVE-3_ManuelClose")
      Visibility <- "HMI_Popup_POPUP{6}"
      on Release: ResetBit("VALVE-H_VALVE-3_ManuelClose")
   Switch "Switch_3" at 189,287 size 130x55; TextOn 'OTO'; CaptionText 'Switch'; TextOff 'MAN'
      Visibility <- "HMI_Popup_POPUP{6}"
   Button "Button_9" at 264,237 size 57x36; TextOff 'Text'; PictureOff "button"
      on Press: InvertBit("HMI_Popup_POPUP{6}")
      Visibility <- "HMI_Popup_POPUP{6}"
   TextField "Text field_5" at 39,242 size 134x33; Text 'VALVE-3'
      Visibility <- "HMI_Popup_POPUP{6}"
   Rectangle "Rectangle_6" at 124,307 size 20x18
      Visibility <- "HMI_Popup_POPUP{6}"
      Appearance <- "VALVE-H_VALVE-3_ValveStatus"
   TextField "Text field_6" at 51,307 size 45x17; Text 'OPENED'
      Visibility <- "HMI_Popup_POPUP{6}"
   Rectangle "Rectangle_7" at 372,227 size 300x170
      Visibility <- "HMI_Popup_POPUP{7}"
   Button "Button_10" at 387,347 size 133x41; TextOn 'AÇILDI'; TextOff 'OPEN'
      on Press: SetBit("VALVE-H_VALVE-4_ManuelOpen")
      Visibility <- "HMI_Popup_POPUP{7}"
      on Release: ResetBit("VALVE-H_VALVE-4_ManuelOpen")
   Button "Button_11" at 525,347 size 133x41; TextOn 'KAPANDI'; TextOff 'CLOSE'
      on Press: SetBit("VALVE-H_VALVE-3_ManuelClose")
      Visibility <- "HMI_Popup_POPUP{7}"
      on Release: ResetBit("VALVE-H_VALVE-3_ManuelClose")
   Switch "Switch_4" at 532,282 size 130x55; TextOn 'OTO'; CaptionText 'Switch'; TextOff 'MAN'
      Visibility <- "HMI_Popup_POPUP{7}"
   Button "Button_12" at 607,232 size 57x36; TextOff 'Text'; PictureOff "button"
      on Press: InvertBit("HMI_Popup_POPUP{7}")
      Visibility <- "HMI_Popup_POPUP{7}"
   TextField "Text field_7" at 382,237 size 134x33; Text 'VALVE-4'
      Visibility <- "HMI_Popup_POPUP{7}"
   Rectangle "Rectangle_8" at 467,302 size 20x18
      Visibility <- "HMI_Popup_POPUP{7}"
      Appearance <- "VALVE-H_VALVE-4_ValveStatus"
   TextField "Text field_8" at 394,302 size 45x17; Text 'OPENED'
      Visibility <- "HMI_Popup_POPUP{7}"
   Group "Group" at 20,20 size 300x170
   Group "Group_1" at 376,20 size 300x170
   Group "Group_2" at 372,227 size 300x170
   Group "Group_3" at 29,232 size 300x170

screen "popup_cvana" 800x480
   Rectangle "Rectangle_1" at 38,239 size 300x170
      Visibility <- "HMI_Popup_POPUP{10}"
   IOField "I/O field_1" at 61,333 size 101x35; FormatPattern 999; Unit  %
      Visibility <- "HMI_Popup_POPUP{10}"
      ProcessValue <- "HMI_CValve-3_Set"
   TextField "Text field_1" at 45,249 size 175x32; Text 'CONTROL VALVE-3'
      Visibility <- "HMI_Popup_POPUP{10}"
   Switch "Switch_1" at 189,321 size 130x55; TextOn 'OTO'; CaptionText 'Switch'; TextOff 'MAN'
      Visibility <- "HMI_Popup_POPUP{10}"
   Button "Button_1" at 274,246 size 57x36; TextOff 'Text'; PictureOff "button"
      on Press: InvertBit("HMI_Popup_POPUP{10}")
      Visibility <- "HMI_Popup_POPUP{10}"
   Rectangle "Rectangle_2" at 402,53 size 300x170
      Visibility <- "HMI_Popup_POPUP{9}"
   IOField "I/O field_2" at 425,147 size 101x35; FormatPattern 999; Unit  %
      Visibility <- "HMI_Popup_POPUP{9}"
      ProcessValue <- "HMI_CValve-2_Set"
   TextField "Text field_2" at 409,63 size 175x32; Text 'CONTROL VALVE-2'
      Visibility <- "HMI_Popup_POPUP{9}"
   Switch "Switch_2" at 553,135 size 130x55; TextOn 'OTO'; CaptionText 'Switch'; TextOff 'MAN'
      Visibility <- "HMI_Popup_POPUP{9}"
   Button "Button_2" at 638,60 size 57x36; TextOff 'Text'; PictureOff "button"
      on Press: InvertBit("HMI_Popup_POPUP{9}")
      Visibility <- "HMI_Popup_POPUP{9}"
   Rectangle "Rectangle_3" at 403,243 size 300x170
      Visibility <- "HMI_Popup_POPUP{11}"
   IOField "I/O field_3" at 426,337 size 101x35; FormatPattern 999; Unit  %
      ProcessValue <- "HMI_CValve-1_Set"
      Visibility <- "HMI_Popup_POPUP{11}"
   TextField "Text field_3" at 410,253 size 175x32; Text 'CONTROL VALVE-4'
      Visibility <- "HMI_Popup_POPUP{11}"
   Switch "Switch_4" at 554,325 size 130x55; TextOn 'OTO'; CaptionText 'Switch'; TextOff 'MAN'
      Visibility <- "HMI_Popup_POPUP{11}"
   Button "Button_3" at 639,250 size 57x36; TextOff 'Text'; PictureOff "button"
      on Press: InvertBit("HMI_Popup_POPUP{11}")
      Visibility <- "HMI_Popup_POPUP{11}"
   Group "Group_1" at 402,53 size 300x170
   Group "Group_2" at 403,243 size 300x170
   Group "Group_3" at 38,239 size 300x170
   Rectangle "Rectangle_30" at 38,53 size 300x170
      Visibility <- "HMI_Popup_POPUP{8}"
   IOField "I/O field_18" at 61,147 size 101x35; FormatPattern 999; Unit  %
      Visibility <- "HMI_Popup_POPUP{8}"
      ProcessValue <- "HMI_CValve-1_Set"
   TextField "Text field_26" at 45,63 size 175x32; Text 'CONTROL VALVE-1'
      Visibility <- "HMI_Popup_POPUP{8}"
   Switch "Switch_3" at 189,135 size 130x55; TextOn 'OTO'; CaptionText 'Switch'; TextOff 'MAN'
      Visibility <- "HMI_Popup_POPUP{8}"
   Button "Button_5" at 274,60 size 57x36; TextOff 'Text'; PictureOff "button"
      on Press: InvertBit("HMI_Popup_POPUP{8}")
      Visibility <- "HMI_Popup_POPUP{8}"
*)